(* Logix 5000 project; controller PLC_MCC1300_75F1 vendor 1 type 14 code 166 rev 32.11; software revision 32.04; part 11 of 83 *)
(* tags used below, declared in another part *)
   CONV1_MS_ACCUM : ALIAS FOR N30[1];
   CONV2_MS_ACCUM : ALIAS FOR N30[2];
   M302SpeedUp : MAC_SpeedUp;
   M310B : MAC_Conveyor;
   M311 : MAC_Conveyor;
   M311A : MAC_Rotator;
   M312 : MAC_Conveyor_Single;
   M315A : MAC_Conveyor;
   M315B : MAC_Conveyor;
   M316 : MAC_Conveyor;
   M316A : MAC_Rotator;
   M317 : MAC_Conveyor_Single;
   M351 : MAC_Conveyor;
   M352 : MAC_Conveyor;
   M353 : MAC_Conveyor;
   O : INT[128];
   TMP_d : DINT;
   TMP_xPositioning : BOOL;
   TMP_xReverse : BOOL;
   TMP_xRun : BOOL;
   xAlwaysOFF : BOOL;
   Z300_Conveyor : UDT_StandConv[29];
   Z300_Conveyor_Conf : UDT_Conveyor_Config[29];

        [14].dWidthConveyor_cmm := 450000, [14].dPitchRoller := 25000, [14].dMachineIndex := 14, [14].dZoneConveyor := 2, [14].dMotorNumber := 1, [14].dSpaceRestartPlate_cmm := 250000, [14].xWaitGlassForStop := 1, [14].rAccH_ms2 := 1.2, [14].rDecH_ms2 := 1.2, [14].rAccH_s := 1.25, [14].rDecH_s := 1.25, [14].rAccL_ms2 := 0.7, [14].rDecL_ms2 := 0.7, [14].rAccL_s := 2.14, [14].rDecL_s := 2.14, [14].rgxAllowedCullet := 16777216, [14].rgxAllowedQuality := 536870912); {access None}
        [7]   // M303M1
        [5]   // M302M6
        [0]   // M302M1
        [10]   // M305M1
        [11]   // M306M1
        [13]   // M307AM2
        [1]   // M302M2
        [2]   // M302M3
        [3]   // M302M4
        [4]   // M302M5
        [6]   // M302M7
        [8]   // M303M2
        [9]   // M304M1
        [28]   // M315M3
        [27]   // M315M2
        [26]   // M315M1
        [25]   // M360M1
        [24]   // M310M3
        [23]   // M310M2
        [22]   // M310M1
        [21]   // M350M1
        [20]   // M307FM1
        [19]   // M307EM1
        [18]   // M307DM1
        [17]   // M307CM1
        [16]   // M30BFM1
        [15]   // M307AM4
        [14]   // M307AM3
        [12]   // M307AM1
   Z300_Conveyor_HMR : MAC_Conveyor_ZC_HMR[29] := ([0].rgdState[0] := 3, [0].rgdState[1] := 1, [1].rgdState[0] := 3, [1].rgdState[1] := 1, [2].rgdState[0] := 3, [2].rgdState[1] := 1, [3].xPlatePresence := 1, [3].rgdState[0] := 3, [3].rgdState[1] := 1, [4].xPlatePresence := 1, [4].rgdState[0] := 3, [4].rgdState[1] := 1, [5].xPlatePresence := 1, [5].rgdState[0] := 3, [5].rgdState[1] := 3, [6].xPlatePresence := 1, [6].rgdState[0] := 3, [6].rgdState[1] := 1, [7].xPlatePresence := 1, [7].rgdState[0] := 3, [7].rgdState[1] := 1, [8].xPlatePresence := 1, [8].rgdState[0] := 3, [8].rgdState[1] := 1, [9].rgdState[0] := 3, [9].rgdState[1] := 1, [10].xPlatePresence := 1, [10].rgdState[0] := 3, [10].rgdState[1] := 1, [11].xPlatePresence := 1, [11].rgdState[0] := 3, [11].rgdState[1] := 3, [12].rgdState[0] := 3, [12].rgdState[1] := 1, [13].xPlatePresence := 1, [13].rgdState[0] := 3, [13].rgdState[1] := 3, [14].rgdState[0] := 3, [14].rgdState[1] := 3); {access Read Only}
        [0]   // M302M1
        [10]   // M305M1
        [21]   // M350M1
        [25]   // M360M1
        [1]   // M302M2
        [2]   // M302M3
        [3]   // M302M4
        [4]   // M302M5
        [8]   // M303M2
        [9]   // M304M1
        [12]   // M307AM1
        [6]   // M302M7
        [7]   // M303M1
        [11]   // M306M1
        [5]   // M302M6
        [13]   // M307AM2
        [14]   // M307AM3
        [15]   // M307AM4
        [16]   // M307BM1
        [17]   // M307CM1
        [18]   // M307DM1
        [19]   // M307EM1
        [20]   // M307FM1
        [22]   // M310BM1
        [23]   // M310BM2
        [24]   // M310BM3
        [26]   // M315BM1
        [27]   // M315BM2
        [28]   // M315BM3
   Z300_Conveyor_HMW : MAC_Conveyor_ZC_HMW[29];
        [5]   // M302M6
        [6]   // M302M7
        [0]   // M302M1
        [10]   // M305M1
        [21]   // M350M1
        [25]   // M360M1
        [1]   // M302M2
        [2]   // M302M3
        [3]   // M302M4
        [4]   // M302M5
        [8]   // M303M2
        [9]   // M304M1
        [7]   // M303M1
        [11]   // M306M1
        [12]   // M307AM1
        [13]   // M307AM2
        [14]   // M307AM3
        [15]   // M307AM4
        [16]   // M307BM1
        [17]   // M307CM1
        [18]   // M307DM1
        [19]   // M307EM1
        [20]   // M307FM1
        [22]   // M310BM1
        [23]   // M310BM2
        [24]   // M310BM3
        [26]   // M315BM1
        [27]   // M315BM2
        [28]   // M315BM3
   Z300_Conveyor_IN_MOTION : MAC_Conveyor_ZC_IN_MOTION[29] := ([0].DR_MAJ_M[0].FLAGS := -1509949438, [0].DR_MAJ_M[0].EN := 1, [0].DR_MAJ_M[0].DN := 1, [0].DR_MAJ_M[0].IP := 1, [0].DR_MAJ_M[0].DECEL := 1, [0].DR_MAM_M[0].FLAGS := 33554432, [0].DR_MRP_M[0].FLAGS := 33554432, [0].DR_MAR_M[0].FLAGS := 33554432, [0].DR_MASall_M[0].FLAGS := 704643072, [0].DR_MASall_M[0].DN := 1, [0].DR_MASall_M[0].PC := 1, [0].DR_MASjog_M[0].FLAGS := 704643072, [0].DR_MASjog_M[0].DN := 1, [0].DR_MASjog_M[0].PC := 1, [0].DR_MASpos_M[0].FLAGS := 33554432, [1].DR_MAJ_M[0].FLAGS := -1509949440, [1].DR_MAJ_M[0].EN := 1, [1].DR_MAJ_M[0].DN := 1, [1].DR_MAJ_M[0].IP := 1, [1].DR_MAM_M[0].FLAGS := 33554432, [1].DR_MRP_M[0].FLAGS := 33554432, [1].DR_MAR_M[0].FLAGS := 33554432, [1].DR_MASall_M[0].FLAGS := 704643072, [1].DR_MASall_M[0].DN := 1, [1].DR_MASall_M[0].PC := 1, [1].DR_MASjog_M[0].FLAGS := 704643072, [1].DR_MASjog_M[0].DN := 1, [1].DR_MASjog_M[0].PC := 1, [1].DR_MASpos_M[0].FLAGS := 33554432, [2].DR_MAJ_M[0].FLAGS := -1509949440, [2].DR_MAJ_M[0].EN := 1, [2].DR_MAJ_M[0].DN := 1, [2].DR_MAJ_M[0].IP := 1, [2].DR_MAM_M[0].FLAGS := 33554432, [2].DR_MASall_M[0].FLAGS := 704643072, [2].DR_MASall_M[0].DN := 1, [2].DR_MASall_M[0].PC := 1, [2].DR_MASjog_M[0].FLAGS := 704643072, [2].DR_MASjog_M[0].DN := 1, [2].DR_MASjog_M[0].PC := 1, [2].DR_MASpos_M[0].FLAGS := 33554432, [3].DR_MAJ_M[0].FLAGS := -1509949440, [3].DR_MAJ_M[0].EN := 1, [3].DR_MAJ_M[0].DN := 1, [3].DR_MAJ_M[0].IP := 1, [3].DR_MAM_M[0].FLAGS := 33554432, [3].DR_MASall_M[0].FLAGS := 704643072, [3].DR_MASall_M[0].DN := 1, [3].DR_MASall_M[0].PC := 1, [3].DR_MASjog_M[0].FLAGS := 704643072, [3].DR_MASjog_M[0].DN := 1, [3].DR_MASjog_M[0].PC := 1, [3].DR_MASpos_M[0].FLAGS := 33554432, [4].DR_MAJ_M[0].FLAGS := -1509949440, [4].DR_MAJ_M[0].EN := 1, [4].DR_MAJ_M[0].DN := 1, [4].DR_MAJ_M[0].IP := 1, [4].DR_MAM_M[0].FLAGS := 33554432, [4].DR_MRP_M[0].FLAGS := 33554432, [4].DR_MAR_M[0].FLAGS := 33554432,
        [4].DR_MASall_M[0].FLAGS := 704643072, [4].DR_MASall_M[0].DN := 1, [4].DR_MASall_M[0].PC := 1, [4].DR_MASjog_M[0].FLAGS := 704643072, [4].DR_MASjog_M[0].DN := 1, [4].DR_MASjog_M[0].PC := 1, [4].DR_MASpos_M[0].FLAGS := 33554432, [5].DR_MAJ_M[0].FLAGS := -1509949440, [5].DR_MAJ_M[0].EN := 1, [5].DR_MAJ_M[0].DN := 1, [5].DR_MAJ_M[0].IP := 1, [5].DR_MAJ_M[1].FLAGS := -1509949440, [5].DR_MAJ_M[1].EN := 1, [5].DR_MAJ_M[1].DN := 1, [5].DR_MAJ_M[1].IP := 1, [5].DR_MAM_M[0].FLAGS := 33554432, [5].DR_MAM_M[1].FLAGS := 33554432, [5].DR_MRP_M[0].FLAGS := 33554432, [5].DR_MRP_M[1].FLAGS := 33554432, [5].DR_MAR_M[0].FLAGS := 33554432, [5].DR_MAR_M[1].FLAGS := 33554432, [5].DR_MASall_M[0].FLAGS := 704643072, [5].DR_MASall_M[0].DN := 1, [5].DR_MASall_M[0].PC := 1, [5].DR_MASall_M[1].FLAGS := 704643072, [5].DR_MASall_M[1].DN := 1, [5].DR_MASall_M[1].PC := 1, [5].DR_MASjog_M[0].FLAGS := 704643072, [5].DR_MASjog_M[0].DN := 1, [5].DR_MASjog_M[0].PC := 1, [5].DR_MASjog_M[1].FLAGS := 704643072, [5].DR_MASjog_M[1].DN := 1, [5].DR_MASjog_M[1].PC := 1, [5].DR_MASpos_M[0].FLAGS := 33554432, [5].DR_MASpos_M[1].FLAGS := 33554432, [6].DR_MAJ_M[0].FLAGS := -1509949440, [6].DR_MAJ_M[0].EN := 1, [6].DR_MAJ_M[0].DN := 1, [6].DR_MAJ_M[0].IP := 1, [6].DR_MAM_M[0].FLAGS := 33554432, [6].DR_MRP_M[0].FLAGS := 33554432, [6].DR_MAR_M[0].FLAGS := 33554432, [6].DR_MASall_M[0].FLAGS := 704643072, [6].DR_MASall_M[0].DN := 1, [6].DR_MASall_M[0].PC := 1, [6].DR_MASjog_M[0].FLAGS := 704643072, [6].DR_MASjog_M[0].DN := 1, [6].DR_MASjog_M[0].PC := 1, [6].DR_MASpos_M[0].FLAGS := 33554432, [7].DR_MAJ_M[0].FLAGS := -1509949440, [7].DR_MAJ_M[0].EN := 1, [7].DR_MAJ_M[0].DN := 1, [7].DR_MAJ_M[0].IP := 1, [7].DR_MAM_M[0].FLAGS := 33554432, [7].DR_MRP_M[0].FLAGS := 33554432, [7].DR_MAR_M[0].FLAGS := 33554432, [7].DR_MASall_M[0].FLAGS := 704643072, [7].DR_MASall_M[0].DN := 1, [7].DR_MASall_M[0].PC := 1, [7].DR_MASjog_M[0].FLAGS := 704643072,
        [7].DR_MASjog_M[0].DN := 1, [7].DR_MASjog_M[0].PC := 1, [7].DR_MASpos_M[0].FLAGS := 33554432, [8].DR_MAJ_M[0].FLAGS := -1509949440, [8].DR_MAJ_M[0].EN := 1, [8].DR_MAJ_M[0].DN := 1, [8].DR_MAJ_M[0].IP := 1, [8].DR_MAM_M[0].FLAGS := 33554432, [8].DR_MASall_M[0].FLAGS := 704643072, [8].DR_MASall_M[0].DN := 1, [8].DR_MASall_M[0].PC := 1, [8].DR_MASjog_M[0].FLAGS := 704643072, [8].DR_MASjog_M[0].DN := 1, [8].DR_MASjog_M[0].PC := 1, [8].DR_MASpos_M[0].FLAGS := 33554432, [9].DR_MAJ_M[0].FLAGS := -1509949440, [9].DR_MAJ_M[0].EN := 1, [9].DR_MAJ_M[0].DN := 1, [9].DR_MAJ_M[0].IP := 1, [9].DR_MAM_M[0].FLAGS := 33554432, [9].DR_MRP_M[0].FLAGS := 33554432, [9].DR_MAR_M[0].FLAGS := 33554432, [9].DR_MASall_M[0].FLAGS := 704643072, [9].DR_MASall_M[0].DN := 1, [9].DR_MASall_M[0].PC := 1, [9].DR_MASjog_M[0].FLAGS := 704643072, [9].DR_MASjog_M[0].DN := 1, [9].DR_MASjog_M[0].PC := 1, [9].DR_MASpos_M[0].FLAGS := 33554432, [10].DR_MAJ_M[0].FLAGS := -1509949440, [10].DR_MAJ_M[0].EN := 1, [10].DR_MAJ_M[0].DN := 1, [10].DR_MAJ_M[0].IP := 1, [10].DR_MAM_M[0].FLAGS := 33554432, [10].DR_MRP_M[0].FLAGS := 33554432, [10].DR_MAR_M[0].FLAGS := 33554432, [10].DR_MASall_M[0].FLAGS := 704643072, [10].DR_MASall_M[0].DN := 1, [10].DR_MASall_M[0].PC := 1, [10].DR_MASjog_M[0].FLAGS := 704643072, [10].DR_MASjog_M[0].DN := 1, [10].DR_MASjog_M[0].PC := 1, [10].DR_MASpos_M[0].FLAGS := 33554432, [11].DR_MAJ_M[0].FLAGS := -1509949440, [11].DR_MAJ_M[0].EN := 1, [11].DR_MAJ_M[0].DN := 1, [11].DR_MAJ_M[0].IP := 1, [11].DR_MAJ_M[1].FLAGS := -1509949440, [11].DR_MAJ_M[1].EN := 1, [11].DR_MAJ_M[1].DN := 1, [11].DR_MAJ_M[1].IP := 1, [11].DR_MAM_M[0].FLAGS := 33554432, [11].DR_MAM_M[1].FLAGS := 33554432, [11].DR_MRP_M[0].FLAGS := 33554432, [11].DR_MRP_M[1].FLAGS := 33554432, [11].DR_MAR_M[0].FLAGS := 33554432, [11].DR_MAR_M[1].FLAGS := 33554432, [11].DR_MASall_M[0].FLAGS := 704643072, [11].DR_MASall_M[0].DN := 1, [11].DR_MASall_M[0].PC := 1,
        [11].DR_MASall_M[1].FLAGS := 704643072, [11].DR_MASall_M[1].DN := 1, [11].DR_MASall_M[1].PC := 1, [11].DR_MASjog_M[0].FLAGS := 704643072, [11].DR_MASjog_M[0].DN := 1, [11].DR_MASjog_M[0].PC := 1, [11].DR_MASjog_M[1].FLAGS := 704643072, [11].DR_MASjog_M[1].DN := 1, [11].DR_MASjog_M[1].PC := 1, [11].DR_MASpos_M[0].FLAGS := 33554432, [11].DR_MASpos_M[1].FLAGS := 33554432, [12].DR_MAJ_M[0].FLAGS := -1509949440, [12].DR_MAJ_M[0].EN := 1, [12].DR_MAJ_M[0].DN := 1, [12].DR_MAJ_M[0].IP := 1, [12].DR_MAM_M[0].FLAGS := 33554432, [12].DR_MRP_M[0].FLAGS := 33554432, [12].DR_MAR_M[0].FLAGS := 33554432, [12].DR_MASall_M[0].FLAGS := 704643072, [12].DR_MASall_M[0].DN := 1, [12].DR_MASall_M[0].PC := 1, [12].DR_MASjog_M[0].FLAGS := 704643072, [12].DR_MASjog_M[0].DN := 1, [12].DR_MASjog_M[0].PC := 1, [12].DR_MASpos_M[0].FLAGS := 33554432, [13].DR_MAJ_M[0].FLAGS := -1509949440, [13].DR_MAJ_M[0].EN := 1, [13].DR_MAJ_M[0].DN := 1, [13].DR_MAJ_M[0].IP := 1, [13].DR_MAJ_M[1].FLAGS := -1509949440, [13].DR_MAJ_M[1].EN := 1, [13].DR_MAJ_M[1].DN := 1, [13].DR_MAJ_M[1].IP := 1, [13].DR_MAM_M[0].FLAGS := 33554432, [13].DR_MAM_M[1].FLAGS := 33554432, [13].DR_MRP_M[0].FLAGS := 33554432, [13].DR_MRP_M[1].FLAGS := 33554432, [13].DR_MAR_M[0].FLAGS := 33554432, [13].DR_MAR_M[1].FLAGS := 33554432, [13].DR_MASall_M[0].FLAGS := 704643072, [13].DR_MASall_M[0].DN := 1, [13].DR_MASall_M[0].PC := 1, [13].DR_MASall_M[1].FLAGS := 704643072, [13].DR_MASall_M[1].DN := 1, [13].DR_MASall_M[1].PC := 1, [13].DR_MASjog_M[0].FLAGS := 704643072, [13].DR_MASjog_M[0].DN := 1, [13].DR_MASjog_M[0].PC := 1, [13].DR_MASjog_M[1].FLAGS := 704643072, [13].DR_MASjog_M[1].DN := 1, [13].DR_MASjog_M[1].PC := 1, [13].DR_MASpos_M[0].FLAGS := 33554432, [13].DR_MASpos_M[1].FLAGS := 33554432, [14].DR_MAJ_M[0].FLAGS := -1509949440, [14].DR_MAJ_M[0].EN := 1, [14].DR_MAJ_M[0].DN := 1, [14].DR_MAJ_M[0].IP := 1, [14].DR_MAJ_M[1].FLAGS := -1509949440, [14].DR_MAJ_M[1].EN := 1, [14].DR_MAJ_M[1].DN := 1,
        [14].DR_MAJ_M[1].IP := 1, [14].DR_MAM_M[0].FLAGS := 33554432, [14].DR_MAM_M[1].FLAGS := 33554432, [14].DR_MRP_M[0].FLAGS := 33554432, [14].DR_MRP_M[1].FLAGS := 33554432, [14].DR_MAR_M[0].FLAGS := 33554432, [14].DR_MAR_M[1].FLAGS := 33554432, [14].DR_MASall_M[0].FLAGS := 704643072, [14].DR_MASall_M[0].DN := 1, [14].DR_MASall_M[0].PC := 1, [14].DR_MASall_M[1].FLAGS := 704643072, [14].DR_MASall_M[1].DN := 1, [14].DR_MASall_M[1].PC := 1, [14].DR_MASjog_M[0].FLAGS := 704643072, [14].DR_MASjog_M[0].DN := 1, [14].DR_MASjog_M[0].PC := 1, [14].DR_MASjog_M[1].FLAGS := 704643072, [14].DR_MASjog_M[1].DN := 1, [14].DR_MASjog_M[1].PC := 1, [14].DR_MASpos_M[0].FLAGS := 33554432, [14].DR_MASpos_M[1].FLAGS := 33554432); {access None}
        [0]   // M302M1
        [10]   // M305M1
        [21]   // M350M1
        [1]   // M302M2
        [2]   // M302M3
        [3]   // M302M4
        [4]   // M302M5
        [8]   // M303M2
        [9]   // M304M1
        [25]   // M360M1
        [5]   // M302M6
        [6]   // M302M7
        [7]   // M303M1
        [11]   // M306M1
        [12]   // M307AM1
        [13]   // M307AM2
        [14]   // M307AM3
        [15]   // M307AM4
        [16]   // M307BM1
        [17]   // M307CM1
        [18]   // M307DM1
        [19]   // M307EM1
        [20]   // M307FM1
        [22]   // M310M1
        [23]   // M310M2
        [24]   // M310M3
        [26]   // M315M1
        [27]   // M315M2
        [28]   // M315M3
   Z300_Conveyor_OUT_MOTION : MAC_Conveyor_ZC_OUT_MOTION[29] := ([0].DR_MSO_M[0].FLAGS := -1610612736, [0].DR_MSO_M[0].EN := 1, [0].DR_MSO_M[0].DN := 1, [0].DR_MSO_M[0].STATE := 1, [0].DR_MSF_M[0].FLAGS := 536870912, [0].DR_MSF_M[0].DN := 1, [0].DR_MSF_M[0].STATUS := 2, [0].DR_MSF_M[0].STATE := 1, [0].DR_MASR_M[0].FLAGS := 570425344, [0].DR_MASR_M[0].DN := 1, [0].DR_MASR_M[0].STATE := 1, [0].DR_MAJ_M[0].FLAGS := -1509949438, [0].DR_MAJ_M[0].EN := 1, [0].DR_MAJ_M[0].DN := 1, [0].DR_MAJ_M[0].IP := 1, [0].DR_MAJ_M[0].DECEL := 1, [0].DR_MAM_M[0].FLAGS := 33554432, [0].DR_MRP_M[0].FLAGS := 33554432, [0].DR_MAR_M[0].FLAGS := 33554432, [0].DR_MDR_M[0].FLAGS := -1845493760, [0].DR_MDR_M[0].EN := 1, [0].DR_MDR_M[0].ER := 1, [0].DR_MDR_M[0].ERR := 11, [0].DR_MCD_M[0].FLAGS := 570425344, [0].DR_MCD_M[0].DN := 1, [0].DR_MCD_M[1].FLAGS := -2147483648, [0].DR_MCD_M[1].EN := 1, [0].DR_MASall_M[0].FLAGS := 704643072, [0].DR_MASall_M[0].DN := 1, [0].DR_MASall_M[0].PC := 1, [0].DR_MASjog_M[0].FLAGS := 704643072, [0].DR_MASjog_M[0].DN := 1, [0].DR_MASjog_M[0].PC := 1, [0].DR_MASpos_M[0].FLAGS := 33554432, [1].DR_MSO_M[0].FLAGS := -1610612736, [1].DR_MSO_M[0].EN := 1, [1].DR_MSO_M[0].DN := 1, [1].DR_MSO_M[0].STATE := 1, [1].DR_MSF_M[0].FLAGS := 570425344, [1].DR_MSF_M[0].DN := 1, [1].DR_MSF_M[0].STATUS := 2, [1].DR_MSF_M[0].STATE := 1, [1].DR_MASR_M[0].FLAGS := 570425344, [1].DR_MASR_M[0].DN := 1, [1].DR_MASR_M[0].STATE := 1, [1].DR_MAJ_M[0].FLAGS := -1509949440, [1].DR_MAJ_M[0].EN := 1, [1].DR_MAJ_M[0].DN := 1, [1].DR_MAJ_M[0].IP := 1, [1].DR_MAM_M[0].FLAGS := 33554432, [1].DR_MRP_M[0].FLAGS := 33554432, [1].DR_MAR_M[0].FLAGS := 33554432, [1].DR_MDR_M[0].FLAGS := -1845493760, [1].DR_MDR_M[0].EN := 1, [1].DR_MDR_M[0].ER := 1, [1].DR_MDR_M[0].ERR := 11, [1].DR_MCD_M[0].FLAGS := 570425344, [1].DR_MCD_M[0].DN := 1, [1].DR_MASall_M[0].FLAGS := 704643072, [1].DR_MASall_M[0].DN := 1,
        [1].DR_MASall_M[0].PC := 1, [1].DR_MASjog_M[0].FLAGS := 704643072, [1].DR_MASjog_M[0].DN := 1, [1].DR_MASjog_M[0].PC := 1, [1].DR_MASpos_M[0].FLAGS := 33554432, [2].DR_MSO_M[0].FLAGS := -1610612736, [2].DR_MSO_M[0].EN := 1, [2].DR_MSO_M[0].DN := 1, [2].DR_MSO_M[0].STATE := 1, [2].DR_MSF_M[0].FLAGS := 570425344, [2].DR_MSF_M[0].DN := 1, [2].DR_MSF_M[0].STATUS := 2, [2].DR_MSF_M[0].STATE := 1, [2].DR_MASR_M[0].FLAGS := 570425344, [2].DR_MASR_M[0].DN := 1, [2].DR_MASR_M[0].STATE := 1, [2].DR_MAJ_M[0].FLAGS := -1509949440, [2].DR_MAJ_M[0].EN := 1, [2].DR_MAJ_M[0].DN := 1, [2].DR_MAJ_M[0].IP := 1, [2].DR_MAM_M[0].FLAGS := 33554432, [2].DR_MRP_M[0].FLAGS := 33554432, [2].DR_MAR_M[0].FLAGS := 33554432, [2].DR_MDR_M[0].FLAGS := -1845493760, [2].DR_MDR_M[0].EN := 1, [2].DR_MDR_M[0].ER := 1, [2].DR_MDR_M[0].ERR := 11, [2].DR_MCD_M[0].FLAGS := 570425344, [2].DR_MCD_M[0].DN := 1, [2].DR_MASall_M[0].FLAGS := 704643072, [2].DR_MASall_M[0].DN := 1, [2].DR_MASall_M[0].PC := 1, [2].DR_MASjog_M[0].FLAGS := 704643072, [2].DR_MASjog_M[0].DN := 1, [2].DR_MASjog_M[0].PC := 1, [2].DR_MASpos_M[0].FLAGS := 33554432, [3].DR_MSO_M[0].FLAGS := -1610612736, [3].DR_MSO_M[0].EN := 1, [3].DR_MSO_M[0].DN := 1, [3].DR_MSO_M[0].STATE := 1, [3].DR_MSF_M[0].FLAGS := 570425344, [3].DR_MSF_M[0].DN := 1, [3].DR_MSF_M[0].STATUS := 2, [3].DR_MSF_M[0].STATE := 1, [3].DR_MASR_M[0].FLAGS := 570425344, [3].DR_MASR_M[0].DN := 1, [3].DR_MASR_M[0].STATE := 1, [3].DR_MAJ_M[0].FLAGS := -1509949440, [3].DR_MAJ_M[0].EN := 1, [3].DR_MAJ_M[0].DN := 1, [3].DR_MAJ_M[0].IP := 1, [3].DR_MAM_M[0].FLAGS := 33554432, [3].DR_MRP_M[0].FLAGS := 33554432, [3].DR_MAR_M[0].FLAGS := 33554432, [3].DR_MDR_M[0].FLAGS := -1845493760, [3].DR_MDR_M[0].EN := 1, [3].DR_MDR_M[0].ER := 1, [3].DR_MDR_M[0].ERR := 11, [3].DR_MCD_M[0].FLAGS := 570425344, [3].DR_MCD_M[0].DN := 1,
        [3].DR_MASall_M[0].FLAGS := 704643072, [3].DR_MASall_M[0].DN := 1, [3].DR_MASall_M[0].PC := 1, [3].DR_MASjog_M[0].FLAGS := 704643072, [3].DR_MASjog_M[0].DN := 1, [3].DR_MASjog_M[0].PC := 1, [3].DR_MASpos_M[0].FLAGS := 33554432, [4].DR_MSO_M[0].FLAGS := -1610612736, [4].DR_MSO_M[0].EN := 1, [4].DR_MSO_M[0].DN := 1, [4].DR_MSO_M[0].STATE := 1, [4].DR_MSF_M[0].FLAGS := 570425344, [4].DR_MSF_M[0].DN := 1, [4].DR_MSF_M[0].STATUS := 2, [4].DR_MSF_M[0].STATE := 1, [4].DR_MASR_M[0].FLAGS := 570425344, [4].DR_MASR_M[0].DN := 1, [4].DR_MASR_M[0].STATE := 1, [4].DR_MAJ_M[0].FLAGS := -1509949440, [4].DR_MAJ_M[0].EN := 1, [4].DR_MAJ_M[0].DN := 1, [4].DR_MAJ_M[0].IP := 1, [4].DR_MAM_M[0].FLAGS := 33554432, [4].DR_MRP_M[0].FLAGS := 33554432, [4].DR_MAR_M[0].FLAGS := 33554432, [4].DR_MDR_M[0].FLAGS := -1845493760, [4].DR_MDR_M[0].EN := 1, [4].DR_MDR_M[0].ER := 1, [4].DR_MDR_M[0].ERR := 11, [4].DR_MCD_M[0].FLAGS := -1577058304, [4].DR_MCD_M[0].EN := 1, [4].DR_MCD_M[0].DN := 1, [4].DR_MASall_M[0].FLAGS := 704643072, [4].DR_MASall_M[0].DN := 1, [4].DR_MASall_M[0].PC := 1, [4].DR_MASjog_M[0].FLAGS := 704643072, [4].DR_MASjog_M[0].DN := 1, [4].DR_MASjog_M[0].PC := 1, [4].DR_MASpos_M[0].FLAGS := 33554432, [5].DR_MSO_M[0].FLAGS := -1610612736, [5].DR_MSO_M[0].EN := 1, [5].DR_MSO_M[0].DN := 1, [5].DR_MSO_M[0].STATE := 1, [5].DR_MSO_M[1].FLAGS := -1610612736, [5].DR_MSO_M[1].EN := 1, [5].DR_MSO_M[1].DN := 1, [5].DR_MSO_M[1].STATE := 1, [5].DR_MSF_M[0].FLAGS := 536870912, [5].DR_MSF_M[0].DN := 1, [5].DR_MSF_M[0].STATUS := 2, [5].DR_MSF_M[0].STATE := 1, [5].DR_MSF_M[1].FLAGS := 536870912, [5].DR_MSF_M[1].DN := 1, [5].DR_MSF_M[1].STATUS := 2, [5].DR_MSF_M[1].STATE := 1, [5].DR_MASR_M[0].FLAGS := 570425344, [5].DR_MASR_M[0].DN := 1, [5].DR_MASR_M[0].STATE := 1, [5].DR_MASR_M[1].FLAGS := 570425344, [5].DR_MASR_M[1].DN := 1,
        [5].DR_MASR_M[1].STATE := 1, [5].DR_MAJ_M[0].FLAGS := -1509949440, [5].DR_MAJ_M[0].EN := 1, [5].DR_MAJ_M[0].DN := 1, [5].DR_MAJ_M[0].IP := 1, [5].DR_MAJ_M[1].FLAGS := -1509949440, [5].DR_MAJ_M[1].EN := 1, [5].DR_MAJ_M[1].DN := 1, [5].DR_MAJ_M[1].IP := 1, [5].DR_MAM_M[0].FLAGS := 33554432, [5].DR_MAM_M[1].FLAGS := 33554432, [5].DR_MRP_M[0].FLAGS := 33554432, [5].DR_MRP_M[1].FLAGS := 33554432, [5].DR_MAR_M[0].FLAGS := 33554432, [5].DR_MAR_M[1].FLAGS := 33554432, [5].DR_MDR_M[0].FLAGS := -1845493760, [5].DR_MDR_M[0].EN := 1, [5].DR_MDR_M[0].ER := 1, [5].DR_MDR_M[0].ERR := 11, [5].DR_MDR_M[1].FLAGS := -1845493760, [5].DR_MDR_M[1].EN := 1, [5].DR_MDR_M[1].ER := 1, [5].DR_MDR_M[1].ERR := 11, [5].DR_MCD_M[0].FLAGS := -1577058304, [5].DR_MCD_M[0].EN := 1, [5].DR_MCD_M[0].DN := 1, [5].DR_MCD_M[1].FLAGS := -1577058304, [5].DR_MCD_M[1].EN := 1, [5].DR_MCD_M[1].DN := 1, [5].DR_MASall_M[0].FLAGS := 704643072, [5].DR_MASall_M[0].DN := 1, [5].DR_MASall_M[0].PC := 1, [5].DR_MASall_M[1].FLAGS := 704643072, [5].DR_MASall_M[1].DN := 1, [5].DR_MASall_M[1].PC := 1, [5].DR_MASjog_M[0].FLAGS := 704643072, [5].DR_MASjog_M[0].DN := 1, [5].DR_MASjog_M[0].PC := 1, [5].DR_MASjog_M[1].FLAGS := 704643072, [5].DR_MASjog_M[1].DN := 1, [5].DR_MASjog_M[1].PC := 1, [5].DR_MASpos_M[0].FLAGS := 33554432, [5].DR_MASpos_M[1].FLAGS := 33554432, [6].DR_MSO_M[0].FLAGS := -1610612736, [6].DR_MSO_M[0].EN := 1, [6].DR_MSO_M[0].DN := 1, [6].DR_MSO_M[0].STATE := 1, [6].DR_MSF_M[0].FLAGS := 570425344, [6].DR_MSF_M[0].DN := 1, [6].DR_MSF_M[0].STATUS := 2, [6].DR_MSF_M[0].STATE := 1, [6].DR_MASR_M[0].FLAGS := 570425344, [6].DR_MASR_M[0].DN := 1, [6].DR_MASR_M[0].STATE := 1, [6].DR_MAJ_M[0].FLAGS := -1509949440, [6].DR_MAJ_M[0].EN := 1, [6].DR_MAJ_M[0].DN := 1, [6].DR_MAJ_M[0].IP := 1, [6].DR_MAM_M[0].FLAGS := 33554432, [6].DR_MRP_M[0].FLAGS := 33554432,
        [6].DR_MAR_M[0].FLAGS := 33554432, [6].DR_MDR_M[0].FLAGS := -1845493760, [6].DR_MDR_M[0].EN := 1, [6].DR_MDR_M[0].ER := 1, [6].DR_MDR_M[0].ERR := 11, [6].DR_MCD_M[0].FLAGS := -1577058304, [6].DR_MCD_M[0].EN := 1, [6].DR_MCD_M[0].DN := 1, [6].DR_MASall_M[0].FLAGS := 704643072, [6].DR_MASall_M[0].DN := 1, [6].DR_MASall_M[0].PC := 1, [6].DR_MASjog_M[0].FLAGS := 704643072, [6].DR_MASjog_M[0].DN := 1, [6].DR_MASjog_M[0].PC := 1, [6].DR_MASpos_M[0].FLAGS := 33554432, [7].DR_MSO_M[0].FLAGS := -1610612736, [7].DR_MSO_M[0].EN := 1, [7].DR_MSO_M[0].DN := 1, [7].DR_MSO_M[0].STATE := 1, [7].DR_MSF_M[0].FLAGS := 536870912, [7].DR_MSF_M[0].DN := 1, [7].DR_MSF_M[0].STATUS := 2, [7].DR_MSF_M[0].STATE := 1, [7].DR_MASR_M[0].FLAGS := 570425344, [7].DR_MASR_M[0].DN := 1, [7].DR_MASR_M[0].STATE := 1, [7].DR_MAJ_M[0].FLAGS := -1509949440, [7].DR_MAJ_M[0].EN := 1, [7].DR_MAJ_M[0].DN := 1, [7].DR_MAJ_M[0].IP := 1, [7].DR_MAM_M[0].FLAGS := 33554432, [7].DR_MRP_M[0].FLAGS := 33554432, [7].DR_MAR_M[0].FLAGS := 33554432, [7].DR_MDR_M[0].FLAGS := -1845493760, [7].DR_MDR_M[0].EN := 1, [7].DR_MDR_M[0].ER := 1, [7].DR_MDR_M[0].ERR := 11, [7].DR_MCD_M[0].FLAGS := -1577058304, [7].DR_MCD_M[0].EN := 1, [7].DR_MCD_M[0].DN := 1, [7].DR_MASall_M[0].FLAGS := 704643072, [7].DR_MASall_M[0].DN := 1, [7].DR_MASall_M[0].PC := 1, [7].DR_MASjog_M[0].FLAGS := 704643072, [7].DR_MASjog_M[0].DN := 1, [7].DR_MASjog_M[0].PC := 1, [7].DR_MASpos_M[0].FLAGS := 33554432, [8].DR_MSO_M[0].FLAGS := -1610612736, [8].DR_MSO_M[0].EN := 1, [8].DR_MSO_M[0].DN := 1, [8].DR_MSO_M[0].STATE := 1, [8].DR_MSF_M[0].FLAGS := 536870912, [8].DR_MSF_M[0].DN := 1, [8].DR_MSF_M[0].STATUS := 2, [8].DR_MSF_M[0].STATE := 1, [8].DR_MASR_M[0].FLAGS := 570425344, [8].DR_MASR_M[0].DN := 1, [8].DR_MASR_M[0].STATE := 1, [8].DR_MAJ_M[0].FLAGS := -1509949440, [8].DR_MAJ_M[0].EN := 1,
        [8].DR_MAJ_M[0].DN := 1, [8].DR_MAJ_M[0].IP := 1, [8].DR_MAM_M[0].FLAGS := 33554432, [8].DR_MRP_M[0].FLAGS := 33554432, [8].DR_MAR_M[0].FLAGS := 33554432, [8].DR_MDR_M[0].FLAGS := -1845493760, [8].DR_MDR_M[0].EN := 1, [8].DR_MDR_M[0].ER := 1, [8].DR_MDR_M[0].ERR := 11, [8].DR_MCD_M[0].FLAGS := 570425344, [8].DR_MCD_M[0].DN := 1, [8].DR_MASall_M[0].FLAGS := 704643072, [8].DR_MASall_M[0].DN := 1, [8].DR_MASall_M[0].PC := 1, [8].DR_MASjog_M[0].FLAGS := 704643072, [8].DR_MASjog_M[0].DN := 1, [8].DR_MASjog_M[0].PC := 1, [8].DR_MASpos_M[0].FLAGS := 33554432, [9].DR_MSO_M[0].FLAGS := -1610612736, [9].DR_MSO_M[0].EN := 1, [9].DR_MSO_M[0].DN := 1, [9].DR_MSO_M[0].STATE := 1, [9].DR_MSF_M[0].FLAGS := 536870912, [9].DR_MSF_M[0].DN := 1, [9].DR_MSF_M[0].STATUS := 2, [9].DR_MSF_M[0].STATE := 1, [9].DR_MASR_M[0].FLAGS := 570425344, [9].DR_MASR_M[0].DN := 1, [9].DR_MASR_M[0].STATE := 1, [9].DR_MAJ_M[0].FLAGS := -1509949440, [9].DR_MAJ_M[0].EN := 1, [9].DR_MAJ_M[0].DN := 1, [9].DR_MAJ_M[0].IP := 1, [9].DR_MAM_M[0].FLAGS := 33554432, [9].DR_MRP_M[0].FLAGS := 33554432, [9].DR_MAR_M[0].FLAGS := 33554432, [9].DR_MDR_M[0].FLAGS := -1845493760, [9].DR_MDR_M[0].EN := 1, [9].DR_MDR_M[0].ER := 1, [9].DR_MDR_M[0].ERR := 11, [9].DR_MCD_M[0].FLAGS := 570425344, [9].DR_MCD_M[0].DN := 1, [9].DR_MASall_M[0].FLAGS := 704643072, [9].DR_MASall_M[0].DN := 1, [9].DR_MASall_M[0].PC := 1, [9].DR_MASjog_M[0].FLAGS := 704643072, [9].DR_MASjog_M[0].DN := 1, [9].DR_MASjog_M[0].PC := 1, [9].DR_MASpos_M[0].FLAGS := 33554432, [10].DR_MSO_M[0].FLAGS := -1610612736, [10].DR_MSO_M[0].EN := 1, [10].DR_MSO_M[0].DN := 1, [10].DR_MSO_M[0].STATE := 1, [10].DR_MSF_M[0].FLAGS := 536870912, [10].DR_MSF_M[0].DN := 1, [10].DR_MSF_M[0].STATUS := 2, [10].DR_MSF_M[0].STATE := 1, [10].DR_MASR_M[0].FLAGS := 570425344, [10].DR_MASR_M[0].DN := 1, [10].DR_MASR_M[0].STATE := 1,
        [10].DR_MAJ_M[0].FLAGS := -1509949440, [10].DR_MAJ_M[0].EN := 1, [10].DR_MAJ_M[0].DN := 1, [10].DR_MAJ_M[0].IP := 1, [10].DR_MAM_M[0].FLAGS := 33554432, [10].DR_MRP_M[0].FLAGS := 33554432, [10].DR_MAR_M[0].FLAGS := 33554432, [10].DR_MDR_M[0].FLAGS := -1845493760, [10].DR_MDR_M[0].EN := 1, [10].DR_MDR_M[0].ER := 1, [10].DR_MDR_M[0].ERR := 11, [10].DR_MCD_M[0].FLAGS := 570425344, [10].DR_MCD_M[0].DN := 1, [10].DR_MASall_M[0].FLAGS := 704643072, [10].DR_MASall_M[0].DN := 1, [10].DR_MASall_M[0].PC := 1, [10].DR_MASjog_M[0].FLAGS := 704643072, [10].DR_MASjog_M[0].DN := 1, [10].DR_MASjog_M[0].PC := 1, [10].DR_MASpos_M[0].FLAGS := 33554432, [11].DR_MSO_M[0].FLAGS := -1610612736, [11].DR_MSO_M[0].EN := 1, [11].DR_MSO_M[0].DN := 1, [11].DR_MSO_M[0].STATE := 1, [11].DR_MSO_M[1].FLAGS := -1610612736, [11].DR_MSO_M[1].EN := 1, [11].DR_MSO_M[1].DN := 1, [11].DR_MSO_M[1].STATE := 1, [11].DR_MSF_M[0].FLAGS := 536870912, [11].DR_MSF_M[0].DN := 1, [11].DR_MSF_M[0].STATUS := 2, [11].DR_MSF_M[0].STATE := 1, [11].DR_MSF_M[1].FLAGS := 570425344, [11].DR_MSF_M[1].DN := 1, [11].DR_MSF_M[1].STATUS := 2, [11].DR_MSF_M[1].STATE := 1, [11].DR_MASR_M[0].FLAGS := 570425344, [11].DR_MASR_M[0].DN := 1, [11].DR_MASR_M[0].STATE := 1, [11].DR_MASR_M[1].FLAGS := 301989888, [11].DR_MASR_M[1].ER := 1, [11].DR_MASR_M[1].ERR := 11, [11].DR_MAJ_M[0].FLAGS := -1509949440, [11].DR_MAJ_M[0].EN := 1, [11].DR_MAJ_M[0].DN := 1, [11].DR_MAJ_M[0].IP := 1, [11].DR_MAJ_M[1].FLAGS := -1509949440, [11].DR_MAJ_M[1].EN := 1, [11].DR_MAJ_M[1].DN := 1, [11].DR_MAJ_M[1].IP := 1, [11].DR_MAM_M[0].FLAGS := 33554432, [11].DR_MAM_M[1].FLAGS := 33554432, [11].DR_MRP_M[0].FLAGS := 33554432, [11].DR_MRP_M[1].FLAGS := 33554432, [11].DR_MAR_M[0].FLAGS := 33554432, [11].DR_MAR_M[1].FLAGS := 33554432, [11].DR_MDR_M[0].FLAGS := -1845493760, [11].DR_MDR_M[0].EN := 1, [11].DR_MDR_M[0].ER := 1, [11].DR_MDR_M[0].ERR := 11,
        [11].DR_MDR_M[1].FLAGS := -1845493760, [11].DR_MDR_M[1].EN := 1, [11].DR_MDR_M[1].ER := 1, [11].DR_MDR_M[1].ERR := 11, [11].DR_MCD_M[0].FLAGS := 570425344, [11].DR_MCD_M[0].DN := 1, [11].DR_MCD_M[1].FLAGS := 570425344, [11].DR_MCD_M[1].DN := 1, [11].DR_MASall_M[0].FLAGS := 704643072, [11].DR_MASall_M[0].DN := 1, [11].DR_MASall_M[0].PC := 1, [11].DR_MASall_M[1].FLAGS := 704643072, [11].DR_MASall_M[1].DN := 1, [11].DR_MASall_M[1].PC := 1, [11].DR_MASjog_M[0].FLAGS := 704643072, [11].DR_MASjog_M[0].DN := 1, [11].DR_MASjog_M[0].PC := 1, [11].DR_MASjog_M[1].FLAGS := 704643072, [11].DR_MASjog_M[1].DN := 1, [11].DR_MASjog_M[1].PC := 1, [11].DR_MASpos_M[0].FLAGS := 33554432, [11].DR_MASpos_M[1].FLAGS := 33554432, [12].DR_MSO_M[0].FLAGS := -1610612736, [12].DR_MSO_M[0].EN := 1, [12].DR_MSO_M[0].DN := 1, [12].DR_MSO_M[0].STATE := 1, [12].DR_MSF_M[0].FLAGS := 536870912, [12].DR_MSF_M[0].DN := 1, [12].DR_MSF_M[0].STATUS := 2, [12].DR_MSF_M[0].STATE := 1, [12].DR_MASR_M[0].FLAGS := 570425344, [12].DR_MASR_M[0].DN := 1, [12].DR_MASR_M[0].STATE := 1, [12].DR_MAJ_M[0].FLAGS := -1509949440, [12].DR_MAJ_M[0].EN := 1, [12].DR_MAJ_M[0].DN := 1, [12].DR_MAJ_M[0].IP := 1, [12].DR_MAM_M[0].FLAGS := 33554432, [12].DR_MRP_M[0].FLAGS := 33554432, [12].DR_MAR_M[0].FLAGS := 33554432, [12].DR_MDR_M[0].FLAGS := -1845493760, [12].DR_MDR_M[0].EN := 1, [12].DR_MDR_M[0].ER := 1, [12].DR_MDR_M[0].ERR := 11, [12].DR_MCD_M[0].FLAGS := 570425344, [12].DR_MCD_M[0].DN := 1, [12].DR_MASall_M[0].FLAGS := 704643072, [12].DR_MASall_M[0].DN := 1, [12].DR_MASall_M[0].PC := 1, [12].DR_MASjog_M[0].FLAGS := 704643072, [12].DR_MASjog_M[0].DN := 1, [12].DR_MASjog_M[0].PC := 1, [12].DR_MASpos_M[0].FLAGS := 33554432, [13].DR_MSO_M[0].FLAGS := -1610612736, [13].DR_MSO_M[0].EN := 1, [13].DR_MSO_M[0].DN := 1, [13].DR_MSO_M[0].STATE := 1, [13].DR_MSO_M[1].FLAGS := -1610612736, [13].DR_MSO_M[1].EN := 1, [13].DR_MSO_M[1].DN := 1,
        [13].DR_MSO_M[1].STATE := 1, [13].DR_MSF_M[0].FLAGS := 536870912, [13].DR_MSF_M[0].DN := 1, [13].DR_MSF_M[0].STATUS := 2, [13].DR_MSF_M[0].STATE := 1, [13].DR_MSF_M[1].FLAGS := 536870912, [13].DR_MSF_M[1].DN := 1, [13].DR_MSF_M[1].STATUS := 2, [13].DR_MSF_M[1].STATE := 1, [13].DR_MASR_M[0].FLAGS := 570425344, [13].DR_MASR_M[0].DN := 1, [13].DR_MASR_M[0].STATE := 1, [13].DR_MASR_M[1].FLAGS := 570425344, [13].DR_MASR_M[1].DN := 1, [13].DR_MASR_M[1].STATE := 1, [13].DR_MAJ_M[0].FLAGS := -1509949440, [13].DR_MAJ_M[0].EN := 1, [13].DR_MAJ_M[0].DN := 1, [13].DR_MAJ_M[0].IP := 1, [13].DR_MAJ_M[1].FLAGS := -1509949440, [13].DR_MAJ_M[1].EN := 1, [13].DR_MAJ_M[1].DN := 1, [13].DR_MAJ_M[1].IP := 1, [13].DR_MAM_M[0].FLAGS := 33554432, [13].DR_MAM_M[1].FLAGS := 33554432, [13].DR_MRP_M[0].FLAGS := 33554432, [13].DR_MRP_M[1].FLAGS := 33554432, [13].DR_MAR_M[0].FLAGS := 33554432, [13].DR_MAR_M[1].FLAGS := 33554432, [13].DR_MDR_M[0].FLAGS := -1845493760, [13].DR_MDR_M[0].EN := 1, [13].DR_MDR_M[0].ER := 1, [13].DR_MDR_M[0].ERR := 11, [13].DR_MDR_M[1].FLAGS := -1845493760, [13].DR_MDR_M[1].EN := 1, [13].DR_MDR_M[1].ER := 1, [13].DR_MDR_M[1].ERR := 11, [13].DR_MCD_M[0].FLAGS := 570425344, [13].DR_MCD_M[0].DN := 1, [13].DR_MCD_M[1].FLAGS := 570425344, [13].DR_MCD_M[1].DN := 1, [13].DR_MASall_M[0].FLAGS := 704643072, [13].DR_MASall_M[0].DN := 1, [13].DR_MASall_M[0].PC := 1, [13].DR_MASall_M[1].FLAGS := 704643072, [13].DR_MASall_M[1].DN := 1, [13].DR_MASall_M[1].PC := 1, [13].DR_MASjog_M[0].FLAGS := 704643072, [13].DR_MASjog_M[0].DN := 1, [13].DR_MASjog_M[0].PC := 1, [13].DR_MASjog_M[1].FLAGS := 704643072, [13].DR_MASjog_M[1].DN := 1, [13].DR_MASjog_M[1].PC := 1, [13].DR_MASpos_M[0].FLAGS := 33554432, [13].DR_MASpos_M[1].FLAGS := 33554432, [14].DR_MSO_M[0].FLAGS := -1610612736, [14].DR_MSO_M[0].EN := 1, [14].DR_MSO_M[0].DN := 1, [14].DR_MSO_M[0].STATE := 1, [14].DR_MSO_M[1].FLAGS := -1610612736,
        [14].DR_MSO_M[1].EN := 1, [14].DR_MSO_M[1].DN := 1, [14].DR_MSO_M[1].STATE := 1, [14].DR_MSF_M[0].FLAGS := 570425344, [14].DR_MSF_M[0].DN := 1, [14].DR_MSF_M[0].STATUS := 2, [14].DR_MSF_M[0].STATE := 1, [14].DR_MSF_M[1].FLAGS := 570425344, [14].DR_MSF_M[1].DN := 1, [14].DR_MSF_M[1].STATUS := 2, [14].DR_MSF_M[1].STATE := 1, [14].DR_MASR_M[0].FLAGS := 570425344, [14].DR_MASR_M[0].DN := 1, [14].DR_MASR_M[0].STATE := 1, [14].DR_MASR_M[1].FLAGS := 570425344, [14].DR_MASR_M[1].DN := 1, [14].DR_MASR_M[1].STATE := 1, [14].DR_MAJ_M[0].FLAGS := -1509949440, [14].DR_MAJ_M[0].EN := 1, [14].DR_MAJ_M[0].DN := 1, [14].DR_MAJ_M[0].IP := 1, [14].DR_MAJ_M[1].FLAGS := -1509949440, [14].DR_MAJ_M[1].EN := 1, [14].DR_MAJ_M[1].DN := 1, [14].DR_MAJ_M[1].IP := 1, [14].DR_MAM_M[0].FLAGS := 33554432, [14].DR_MAM_M[1].FLAGS := 33554432, [14].DR_MRP_M[0].FLAGS := 33554432, [14].DR_MRP_M[1].FLAGS := 33554432, [14].DR_MAR_M[0].FLAGS := 33554432, [14].DR_MAR_M[1].FLAGS := 33554432, [14].DR_MDR_M[0].FLAGS := -1845493760, [14].DR_MDR_M[0].EN := 1, [14].DR_MDR_M[0].ER := 1, [14].DR_MDR_M[0].ERR := 11, [14].DR_MDR_M[1].FLAGS := -1845493760, [14].DR_MDR_M[1].EN := 1, [14].DR_MDR_M[1].ER := 1, [14].DR_MDR_M[1].ERR := 11, [14].DR_MCD_M[0].FLAGS := 570425344, [14].DR_MCD_M[0].DN := 1, [14].DR_MCD_M[1].FLAGS := 570425344, [14].DR_MCD_M[1].DN := 1, [14].DR_MASall_M[0].FLAGS := 704643072, [14].DR_MASall_M[0].DN := 1, [14].DR_MASall_M[0].PC := 1, [14].DR_MASall_M[1].FLAGS := 704643072, [14].DR_MASall_M[1].DN := 1, [14].DR_MASall_M[1].PC := 1, [14].DR_MASjog_M[0].FLAGS := 704643072, [14].DR_MASjog_M[0].DN := 1, [14].DR_MASjog_M[0].PC := 1, [14].DR_MASjog_M[1].FLAGS := 704643072, [14].DR_MASjog_M[1].DN := 1, [14].DR_MASjog_M[1].PC := 1, [14].DR_MASpos_M[0].FLAGS := 33554432, [14].DR_MASpos_M[1].FLAGS := 33554432); {access None}
        [5]   // M302M6
        [6]   // M302M7
        [11]   // M306M1
        [0]   // M302M1
        [10]   // M305M1
        [7]   // M303M1
        [21]   // M350M1
        [1]   // M302M2
        [2]   // M302M3
        [3]   // M302M4
        [4]   // M302M5
        [8]   // M303M2
        [9]   // M304M1
        [12]   // M307AM1
        [13]   // M307AM2
        [14]   // M307AM3
        [15]   // M307AM4
        [16]   // M307BM1
        [17]   // M307CM1
        [18]   // M307DM1
        [19]   // M307EM1
        [20]   // M307FM1
        [25]   // M360M1
        [22]   // M310M1
        [23]   // M310M2
        [24]   // M310M3
        [26]   // M315M1
        [27]   // M315M2
        [28]   // M315M3
   Z300_dEndTrackingPosition : DINT := 5395000; {access None}
   Z300_dStartTrackingPosition : DINT; {access None}
   Z300_LineTracking : UDT_LINE_TRACKING := (rgtTrkConv[0].dEndPosition_cmm := 37500, rgtTrkConv[0].dStepAdv_cmm[0] := 679, rgtTrkConv[0].dActualRamp_cmm[0] := 4700, rgtTrkConv[0].dLengthConveyor := 37500, rgtTrkConv[1].dStartPosition_cmm := 37500, rgtTrkConv[1].dEndPosition_cmm := 87500, rgtTrkConv[1].dStepAdv_cmm[0] := 679, rgtTrkConv[1].dActualRamp_cmm[0] := 4700, rgtTrkConv[1].dLengthConveyor := 50000, rgtTrkConv[2].xGlassPresence := 1, rgtTrkConv[2].xPlatePassageNext := 1, rgtTrkConv[2].xGlassPresCom := 1, rgtTrkConv[2].dStartPosition_cmm := 87500, rgtTrkConv[2].dEndPosition_cmm := 212500, rgtTrkConv[2].dStepAdv_cmm[0] := 1800, rgtTrkConv[2].dActualRamp_cmm[0] := 33700, rgtTrkConv[2].dLengthConveyor := 125000, rgtTrkConv[2].dTailPosition_cmm := 179869, rgtTrkConv[2].dIndexCaps := 1, rgtTrkConv[2].Cap[0].xTail := 1, rgtTrkConv[2].Cap[0].xPresence := 1, rgtTrkConv[2].Cap[0].dPointer := 4, rgtTrkConv[2].Cap[0].dTailPos_cmm := 179869, rgtTrkConv[2].Cap[0].dTailPosConv_cmm := 92369, rgtTrkConv[2].Cap[0].dPresenceHead_cmm := 347569, rgtTrkConv[2].Cap[0].dPresenceTail_cmm := 179869, rgtTrkConv[3].xGlassPresence := 1, rgtTrkConv[3].xPlatePassagePrevious := 1, rgtTrkConv[3].xGlassPresCom := 1, rgtTrkConv[3].xHeadPresenceConv := 1, rgtTrkConv[3].dStartPosition_cmm := 212500, rgtTrkConv[3].dEndPosition_cmm := 462500, rgtTrkConv[3].dStepAdv_cmm[0] := 1800, rgtTrkConv[3].dActualRamp_cmm[0] := 33700, rgtTrkConv[3].dLengthConveyor := 250000, rgtTrkConv[3].dHeadPosition_cmm := 349549, rgtTrkConv[3].dIndexCaps := 1, rgtTrkConv[3].Cap[0].xHead := 1, rgtTrkConv[3].Cap[0].xCenter := 1, rgtTrkConv[3].Cap[0].xPresence := 1, rgtTrkConv[3].Cap[0].dPointer := 4, rgtTrkConv[3].Cap[0].dCenterPos_cmm := 265699, rgtTrkConv[3].Cap[0].dCenterPosConv_cmm := 53199, rgtTrkConv[3].Cap[0].dHeadPos_cmm := 349549, rgtTrkConv[3].Cap[0].dHeadPosConv_cmm := 137049, rgtTrkConv[3].Cap[0].dPresenceHead_cmm := 349549, rgtTrkConv[3].Cap[0].dPresenceTail_cmm := 181849, rgtTrkConv[4].xGlassPresence := 1, rgtTrkConv[4].xPlatePassageNext := 1, rgtTrkConv[4].xGlassPresCom := 1, rgtTrkConv[4].dStartPosition_cmm := 462500, rgtTrkConv[4].dEndPosition_cmm := 712500, rgtTrkConv[4].dStepAdv_cmm[0] := 1980, rgtTrkConv[4].dActualRamp_cmm[0] := 33700, rgtTrkConv[4].dLengthConveyor := 250000, rgtTrkConv[4].dTailPosition_cmm := 613600, rgtTrkConv[4].dIndexCaps := 1, rgtTrkConv[4].Cap[0].xTail := 1, rgtTrkConv[4].Cap[0].xPresence := 1, rgtTrkConv[4].Cap[0].dPointer := 2,
        rgtTrkConv[4].Cap[0].dTailPos_cmm := 613600, rgtTrkConv[4].Cap[0].dTailPosConv_cmm := 151100, rgtTrkConv[4].Cap[0].dPresenceHead_cmm := 873600, rgtTrkConv[4].Cap[0].dPresenceTail_cmm := 613600, rgtTrkConv[5].xGlassPresence := 1, rgtTrkConv[5].xPlatePassagePrevious := 1, rgtTrkConv[5].xGlassPresCom := 1, rgtTrkConv[5].xHeadPresenceConv := 1, rgtTrkConv[5].dStartPosition_cmm := 712500, rgtTrkConv[5].dEndPosition_cmm := 1627000, rgtTrkConv[5].dStepAdv_cmm[0] := 1980, rgtTrkConv[5].dStepAdv_cmm[1] := 1980, rgtTrkConv[5].dActualRamp_cmm[0] := 33700, rgtTrkConv[5].dActualRamp_cmm[1] := 33700, rgtTrkConv[5].dLengthConveyor := 914500, rgtTrkConv[5].dHeadPosition_cmm := 1474980, rgtTrkConv[5].dTailPosition_cmm := 1307280, rgtTrkConv[5].dIndexCaps := 2, rgtTrkConv[5].Cap[0].xHead := 1, rgtTrkConv[5].Cap[0].xCenter := 1, rgtTrkConv[5].Cap[0].xPresence := 1, rgtTrkConv[5].Cap[0].dPointer := 2, rgtTrkConv[5].Cap[0].dCenterPos_cmm := 743600, rgtTrkConv[5].Cap[0].dCenterPosConv_cmm := 31100, rgtTrkConv[5].Cap[0].dHeadPos_cmm := 873600, rgtTrkConv[5].Cap[0].dHeadPosConv_cmm := 161100, rgtTrkConv[5].Cap[0].dPresenceHead_cmm := 873600, rgtTrkConv[5].Cap[0].dPresenceTail_cmm := 613600, rgtTrkConv[5].Cap[1].xHead := 1, rgtTrkConv[5].Cap[1].xCenter := 1, rgtTrkConv[5].Cap[1].xTail := 1, rgtTrkConv[5].Cap[1].xPresence := 1, rgtTrkConv[5].Cap[1].dPointer := 7, rgtTrkConv[5].Cap[1].dTailPos_cmm := 1307280, rgtTrkConv[5].Cap[1].dTailPosConv_cmm := 594780, rgtTrkConv[5].Cap[1].dCenterPos_cmm := 1391130, rgtTrkConv[5].Cap[1].dCenterPosConv_cmm := 678630, rgtTrkConv[5].Cap[1].dHeadPos_cmm := 1474980, rgtTrkConv[5].Cap[1].dHeadPosConv_cmm := 762480, rgtTrkConv[5].Cap[1].dPresenceHead_cmm := 1474980, rgtTrkConv[5].Cap[1].dPresenceTail_cmm := 1307280, rgtTrkConv[6].xGlassPresence := 1, rgtTrkConv[6].xGlassPresCom := 1, rgtTrkConv[6].xHeadPresenceConv := 1, rgtTrkConv[6].dStartPosition_cmm := 1627000, rgtTrkConv[6].dEndPosition_cmm := 2127000, rgtTrkConv[6].dStepAdv_cmm[0] := 1980, rgtTrkConv[6].dActualRamp_cmm[0] := 33700, rgtTrkConv[6].dLengthConveyor := 500000, rgtTrkConv[6].dHeadPosition_cmm := 2014180, rgtTrkConv[6].dTailPosition_cmm := 1754180, rgtTrkConv[6].dIndexCaps := 1, rgtTrkConv[6].Cap[0].xHead := 1, rgtTrkConv[6].Cap[0].xCenter := 1, rgtTrkConv[6].Cap[0].xTail := 1, rgtTrkConv[6].Cap[0].xPresence := 1, rgtTrkConv[6].Cap[0].dPointer := 6, rgtTrkConv[6].Cap[0].dTailPos_cmm := 1755800, rgtTrkConv[6].Cap[0].dTailPosConv_cmm := 128800, rgtTrkConv[6].Cap[0].dCenterPos_cmm := 1885800,